(* Logix 5000 project; controller PLC_MCC1300_75F1 vendor 1 type 14 code 166 rev 32.11; software revision 32.04; part 22 of 83 *)
(* tags used below, declared in another part *)
   CM_LineToConveyorStacker_JS1 : CM_LineToConveyorStacker;
   GP_OB_InitializeMain : GP_OB_Initialize;
   M312 : MAC_Conveyor_Single;
   M312_Data : UDT_Convoy_SL;
   M312_HMW : MAC_Conveyor_HMW;
   M312_M3_ChangeSpeed : BOOL;
   M312_M3_DR_IN_MAJ : MOTION_INSTRUCTION;
   M312_M3_DR_L : AXIS_CIP_DRIVE;
   M312_M3_DR_OUT_MAJ : MOTION_INSTRUCTION;
   M312_M3_DR_OUT_MAS : MOTION_INSTRUCTION;
   M312_M3_DR_OUT_MCD : MOTION_INSTRUCTION;
   M312_SpaceConv_Utilities : SpaceConv_Utilities;
   M315_M4_DR_B1 : AXIS_CIP_DRIVE;
   M315A : MAC_Conveyor;
   M315A_ALM : MAC_Conveyor_ALM;
   M315A_Data : UDT_Convoy_SL;
   M315A_HMR : MAC_Conveyor_HMR;
   M315A_HMW : MAC_Conveyor_HMW;
   M315A_M1_DR : AXIS_CIP_DRIVE;
   M315A_M1_DR_IN_MAJ : MOTION_INSTRUCTION;
   M315A_M1_DR_IN_MAR : MOTION_INSTRUCTION;
   M315A_M1_DR_IN_MAS : MOTION_INSTRUCTION;
   M315A_M1_DR_IN_MRP : MOTION_INSTRUCTION;
   M315A_M1_DR_MAFR : MOTION_INSTRUCTION;
   M315A_M1_DR_MDR : MOTION_INSTRUCTION;
   M315A_M1_DR_MSF : MOTION_INSTRUCTION;
   M315A_M1_DR_MSO : MOTION_INSTRUCTION;
   M315A_M1_DR_OUT_MAJ : MOTION_INSTRUCTION;
   M315A_M1_DR_OUT_MAM : MOTION_INSTRUCTION;
   M315A_M1_DR_OUT_MAR : MOTION_INSTRUCTION;
   M315A_M1_DR_OUT_MAS : MOTION_INSTRUCTION;
   M315A_M1_DR_OUT_MCD : MOTION_INSTRUCTION;
   M315A_M1_DR_OUT_MRP : MOTION_INSTRUCTION;
   M315A_SpaceConv_Utilities : SpaceConv_Utilities;
   M315B : MAC_Conveyor;
   M315B_ALM : MAC_Conveyor_ALM;
   M315B_HMR : MAC_Conveyor_HMR;
   M315B_HMW : MAC_Conveyor_HMW;
   M315B_M1_DR_MAFR : MOTION_INSTRUCTION;
   M315B_M1_DR_MSF : MOTION_INSTRUCTION;
   M315B_M1_DR_MSO : MOTION_INSTRUCTION;
   M315B_M1_DR_OUT_MAR : MOTION_INSTRUCTION;
   M315B_M1_DR_OUT_MRP : MOTION_INSTRUCTION;
   M316 : MAC_Conveyor;
   TMP_dDirection : DINT;
   TMP_r : REAL;
   TMP_rAcc : REAL;
   TMP_rDec : REAL;
   TMP_rSpeed : REAL;
   TMP_rTarget_M1 : REAL;
   TMP_xForwardCommadnForCleaningZone : BOOL;
   TMP_xPositioning_M1 : BOOL;
   TMP_xPositioning_M2 : BOOL;
   TMP_xPositioning_M3 : BOOL;
   TMP_xPowerSaving : BOOL;
   TMP_xReverse_M1 : BOOL;
   TMP_xReverse_M2 : BOOL;
   TMP_xReverse_M3 : BOOL;
   TMP_xRun_M1 : BOOL;
   TMP_xRun_M2 : BOOL;
   TMP_xRun_M3 : BOOL;
   xAlwaysOFF : BOOL;
   xAlwaysON : BOOL;
   xDebugOFF : BOOL;
   Z401 : MAC_Zone;
   Z402 : MAC_Zone;
   Z402_HMW : MAC_Zone_HMW;
(* CommandLogic, continued *)

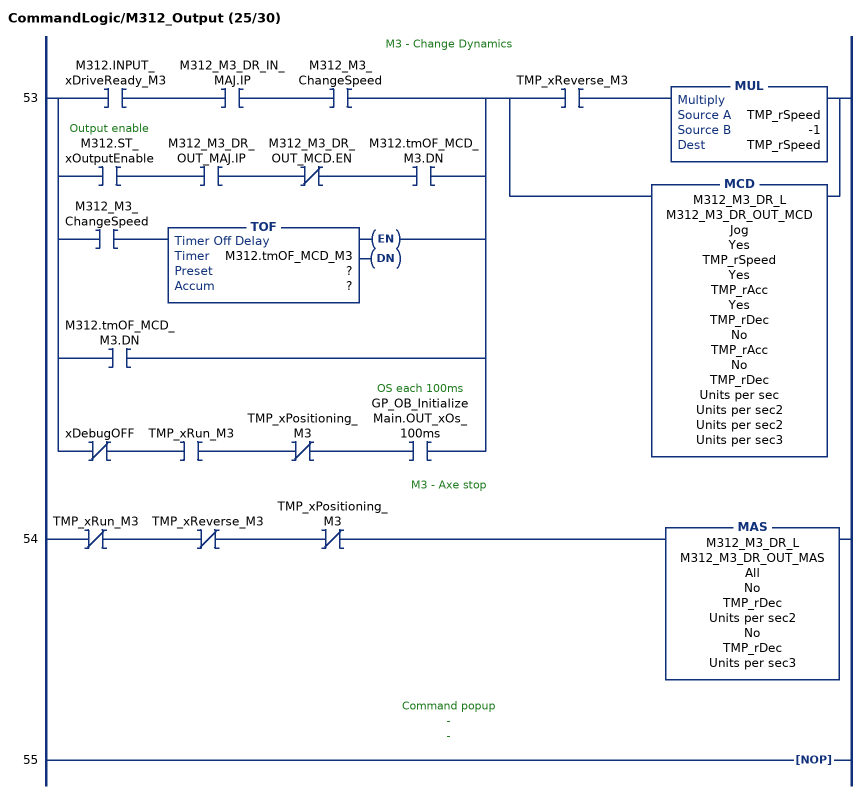
   [picture p215: CommandLogic/M312_Output rungs 53-55]
   // M3 - Change Dynamics
   53: [XIC(M312.INPUT_xDriveReady_M3) XIC(M312_M3_DR_IN_MAJ.IP) XIC(M312_M3_ChangeSpeed) ,XIC(M312.ST_xOutputEnable) XIC(M312_M3_DR_OUT_MAJ.IP) XIO(M312_M3_DR_OUT_MCD.EN) XIC(M312.tmOF_MCD_M3.DN) ,[XIC(M312_M3_ChangeSpeed) TOF(M312.tmOF_MCD_M3,?,?) ,XIC(M312.tmOF_MCD_M3.DN) ] ,XIO(xDebugOFF) XIC(TMP_xRun_M3) XIO(TMP_xPositioning_M3) XIC(GP_OB_InitializeMain.OUT_xOs_100ms) ][XIC(TMP_xReverse_M3) MUL(TMP_rSpeed,-1,TMP_rSpeed) ,MCD(M312_M3_DR_L,M312_M3_DR_OUT_MCD,Jog,Yes,TMP_rSpeed,Yes,TMP_rAcc,Yes,TMP_rDec,No,TMP_rAcc,No,TMP_rDec,Units per sec,Units per sec2,Units per sec2,Units per sec3) ];
   // M3 - Axe stop
   54: XIO(TMP_xRun_M3)XIO(TMP_xReverse_M3)XIO(TMP_xPositioning_M3)MAS(M312_M3_DR_L,M312_M3_DR_OUT_MAS,All,No,TMP_rDec,Units per sec2,No,TMP_rDec,Units per sec3);
   // Command popup
   // -
   // -
   55: NOP();
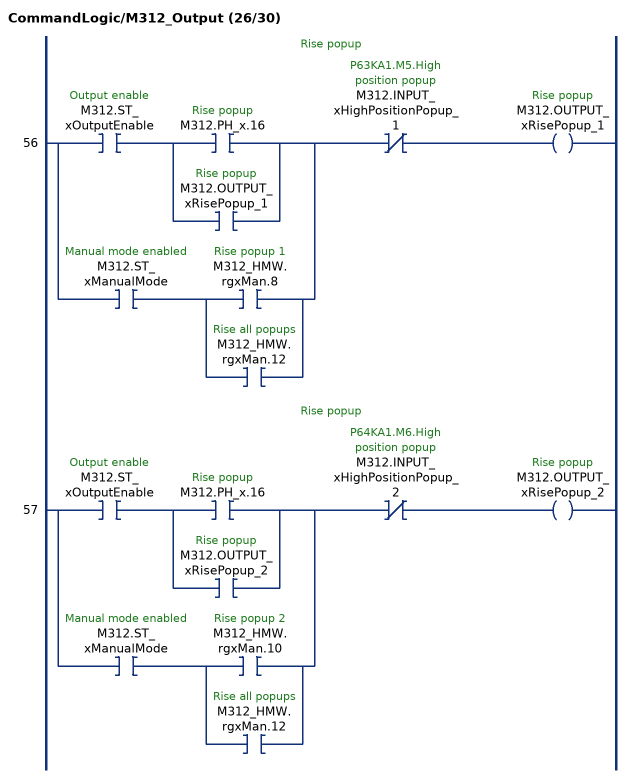
   // Rise popup
   56: [XIC(M312.ST_xOutputEnable) [XIC(M312.PH_x.16) ,XIC(M312.OUTPUT_xRisePopup_1) ] ,XIC(M312.ST_xManualMode) [XIC(M312_HMW.rgxMan.8) ,XIC(M312_HMW.rgxMan.12) ] ]XIO(M312.INPUT_xHighPositionPopup_1)OTE(M312.OUTPUT_xRisePopup_1);
   // Rise popup
   57: [XIC(M312.ST_xOutputEnable) [XIC(M312.PH_x.16) ,XIC(M312.OUTPUT_xRisePopup_2) ] ,XIC(M312.ST_xManualMode) [XIC(M312_HMW.rgxMan.10) ,XIC(M312_HMW.rgxMan.12) ] ]XIO(M312.INPUT_xHighPositionPopup_2)OTE(M312.OUTPUT_xRisePopup_2);
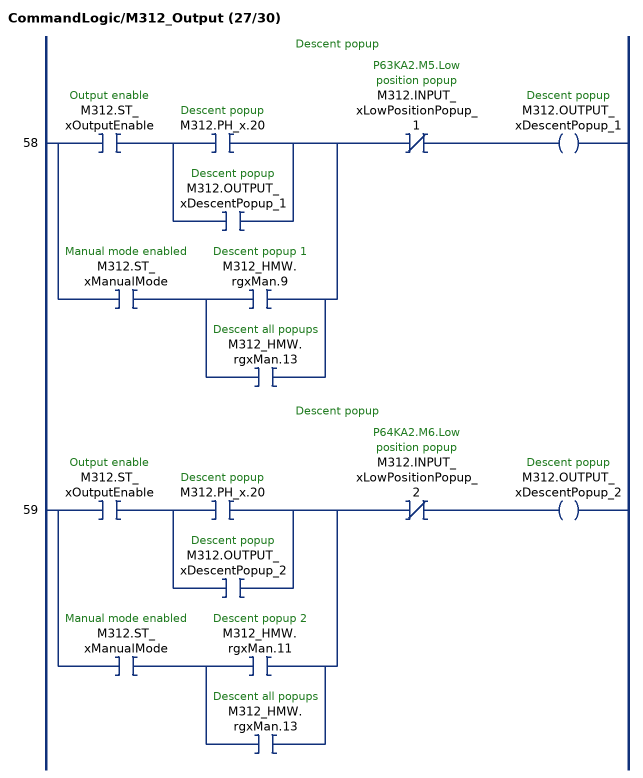
   // Descent popup
   58: [XIC(M312.ST_xOutputEnable) [XIC(M312.PH_x.20) ,XIC(M312.OUTPUT_xDescentPopup_1) ] ,XIC(M312.ST_xManualMode) [XIC(M312_HMW.rgxMan.9) ,XIC(M312_HMW.rgxMan.13) ] ]XIO(M312.INPUT_xLowPositionPopup_1)OTE(M312.OUTPUT_xDescentPopup_1);
   // Descent popup
   59: [XIC(M312.ST_xOutputEnable) [XIC(M312.PH_x.20) ,XIC(M312.OUTPUT_xDescentPopup_2) ] ,XIC(M312.ST_xManualMode) [XIC(M312_HMW.rgxMan.11) ,XIC(M312_HMW.rgxMan.13) ] ]XIO(M312.INPUT_xLowPositionPopup_2)OTE(M312.OUTPUT_xDescentPopup_2);
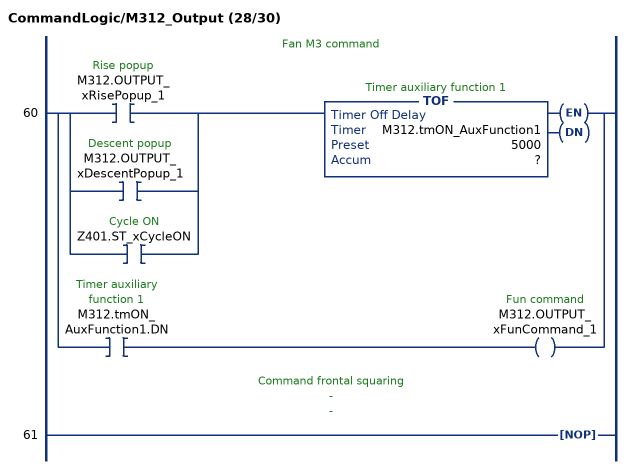
   // Fan M3 command
   60: [[XIC(M312.OUTPUT_xRisePopup_1) ,[XIC(M312.OUTPUT_xDescentPopup_1) ,XIC(Z401.ST_xCycleON) ] ] TOF(M312.tmON_AuxFunction1,?,?) ,XIC(M312.tmON_AuxFunction1.DN) OTE(M312.OUTPUT_xFunCommand_1) ];
   // Command frontal squaring
   // -
   // -
   61: NOP();
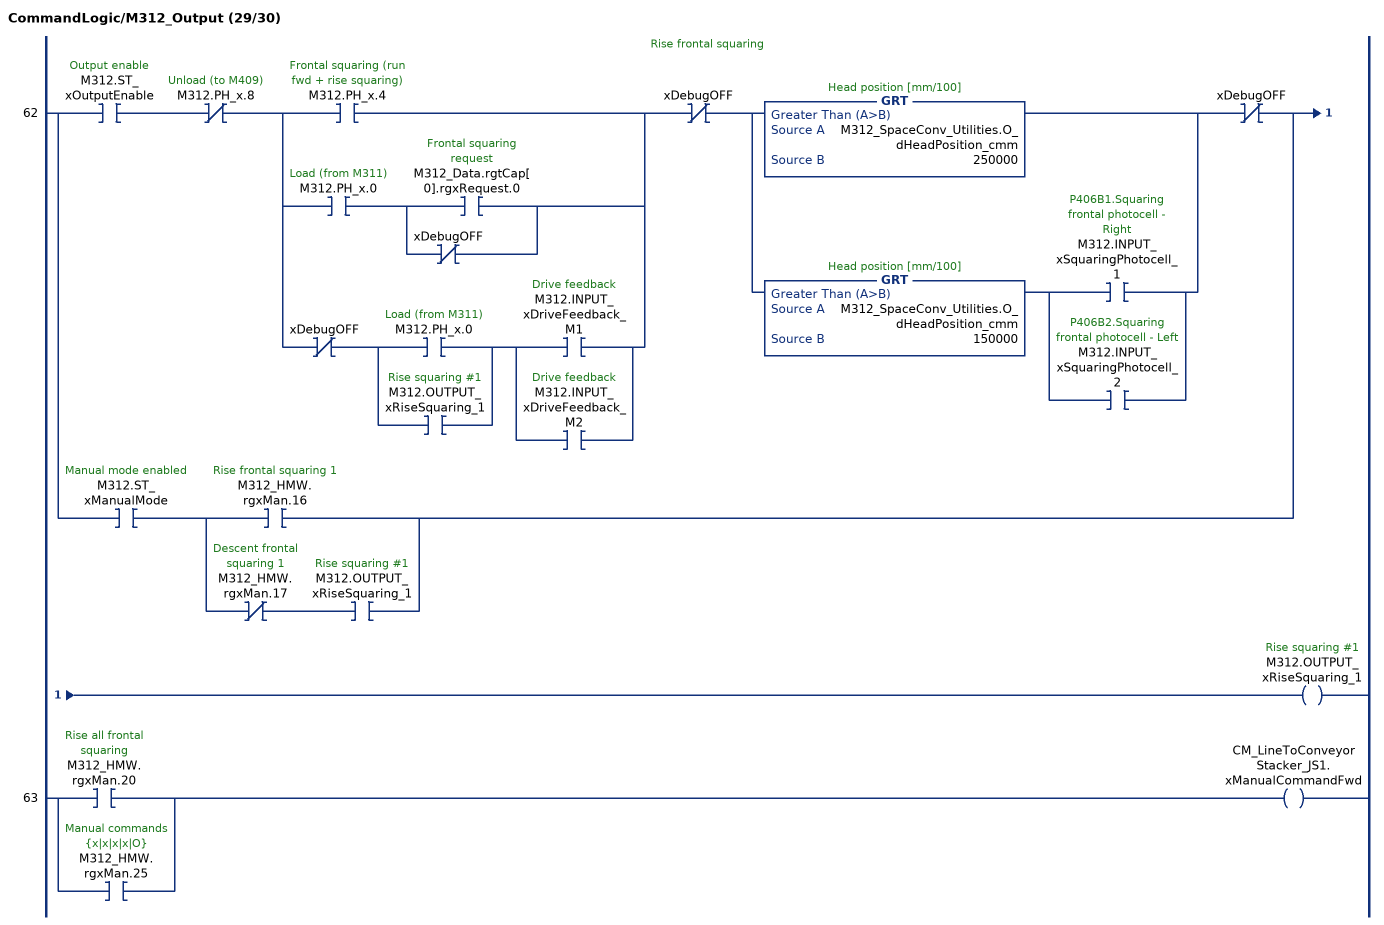
   // Rise frontal squaring
   62: [XIC(M312.ST_xOutputEnable) XIO(M312.PH_x.8) [XIC(M312.PH_x.4) ,XIC(M312.PH_x.0) [XIC(M312_Data.rgtCap[0].rgxRequest.0) ,XIO(xDebugOFF) ] ,XIO(xDebugOFF) [XIC(M312.PH_x.0) ,XIC(M312.OUTPUT_xRiseSquaring_1) ] [XIC(M312.INPUT_xDriveFeedback_M1) ,XIC(M312.INPUT_xDriveFeedback_M2) ] ] XIO(xDebugOFF) [GRT(M312_SpaceConv_Utilities.O_dHeadPosition_cmm,250000) ,GRT(M312_SpaceConv_Utilities.O_dHeadPosition_cmm,150000) [XIC(M312.INPUT_xSquaringPhotocell_1) ,XIC(M312.INPUT_xSquaringPhotocell_2) ] ] XIO(xDebugOFF) ,XIC(M312.ST_xManualMode) [XIC(M312_HMW.rgxMan.16) ,XIO(M312_HMW.rgxMan.17) XIC(M312.OUTPUT_xRiseSquaring_1) ] ]OTE(M312.OUTPUT_xRiseSquaring_1);
   63: [XIC(M312_HMW.rgxMan.20) ,XIC(M312_HMW.rgxMan.25) ]OTE(CM_LineToConveyorStacker_JS1.xManualCommandFwd);
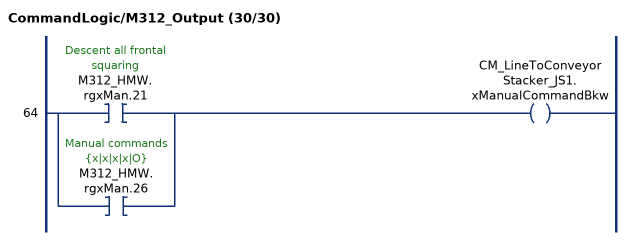
   64: [XIC(M312_HMW.rgxMan.21) ,XIC(M312_HMW.rgxMan.26) ]OTE(CM_LineToConveyorStacker_JS1.xManualCommandBkw);
END_ROUTINE

ROUTINE M315A_Output   (* ladder *)
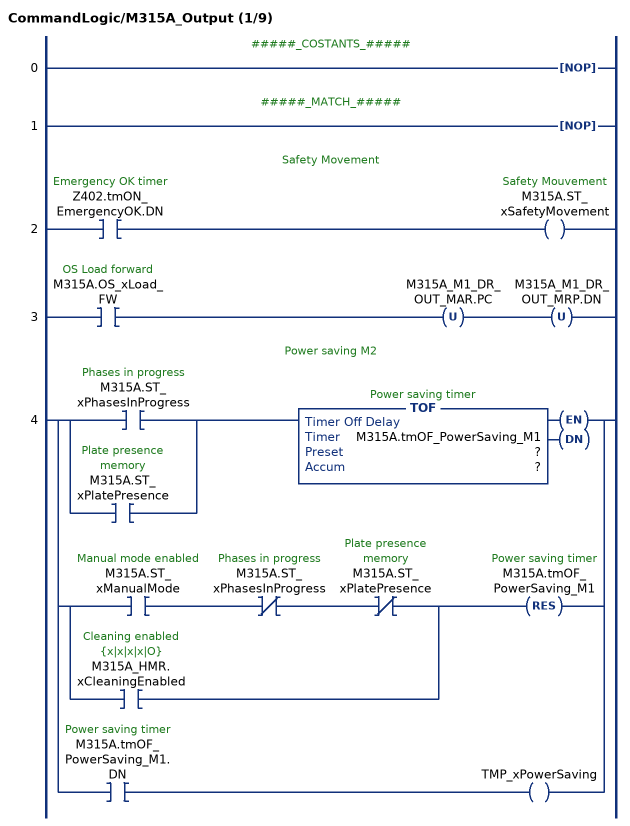
   // #####_COSTANTS_#####
   0: NOP();
   // #####_MATCH_#####
   1: NOP();
   // Safety Movement
   2: XIC(Z402.tmON_EmergencyOK.DN)OTE(M315A.ST_xSafetyMovement);
   3: XIC(M315A.OS_xLoad_FW)OTU(M315A_M1_DR_OUT_MAR.PC)OTU(M315A_M1_DR_OUT_MRP.DN);
   // Power saving M2
   4: [[XIC(M315A.ST_xPhasesInProgress) ,XIC(M315A.ST_xPlatePresence) ] TOF(M315A.tmOF_PowerSaving_M1,?,?) ,[XIC(M315A.ST_xManualMode) XIO(M315A.ST_xPhasesInProgress) XIO(M315A.ST_xPlatePresence) ,XIC(M315A_HMR.xCleaningEnabled) ] RES(M315A.tmOF_PowerSaving_M1) ,XIC(M315A.tmOF_PowerSaving_M1.DN) OTE(TMP_xPowerSaving) ];
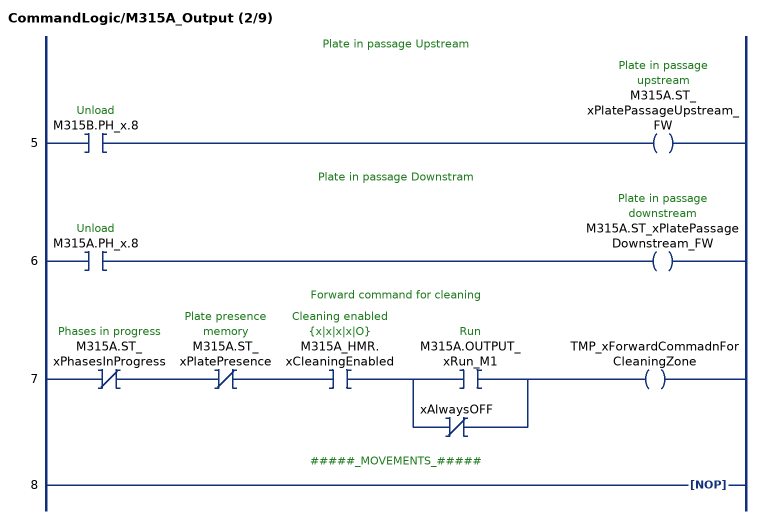
   // Plate in passage Upstream
   5: XIC(M315B.PH_x.8)OTE(M315A.ST_xPlatePassageUpstream_FW);
   // Plate in passage Downstram
   6: XIC(M315A.PH_x.8)OTE(M315A.ST_xPlatePassageDownstream_FW);
   // Forward command for cleaning
   7: XIO(M315A.ST_xPhasesInProgress)XIO(M315A.ST_xPlatePresence)XIC(M315A_HMR.xCleaningEnabled)[XIC(M315A.OUTPUT_xRun_M1) ,XIO(xAlwaysOFF) ]OTE(TMP_xForwardCommadnForCleaningZone);
   // #####_MOVEMENTS_#####
   8: NOP();
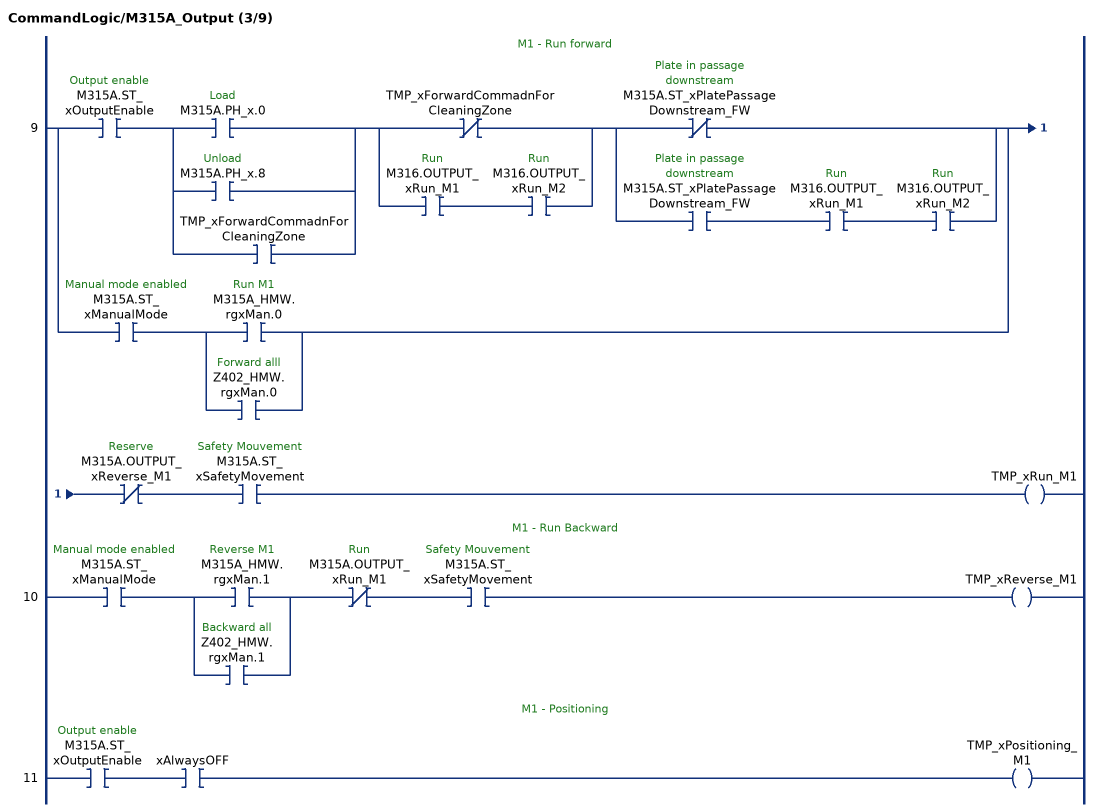
   // M1 - Run forward
   9: [XIC(M315A.ST_xOutputEnable) [XIC(M315A.PH_x.0) ,XIC(M315A.PH_x.8) ,XIC(TMP_xForwardCommadnForCleaningZone) ] [XIO(TMP_xForwardCommadnForCleaningZone) ,XIC(M316.OUTPUT_xRun_M1) XIC(M316.OUTPUT_xRun_M2) ] [XIO(M315A.ST_xPlatePassageDownstream_FW) ,XIC(M315A.ST_xPlatePassageDownstream_FW) XIC(M316.OUTPUT_xRun_M1) XIC(M316.OUTPUT_xRun_M2) ] ,XIC(M315A.ST_xManualMode) [XIC(M315A_HMW.rgxMan.0) ,XIC(Z402_HMW.rgxMan.0) ] ]XIO(M315A.OUTPUT_xReverse_M1)XIC(M315A.ST_xSafetyMovement)OTE(TMP_xRun_M1);
   // M1 - Run Backward
   10: XIC(M315A.ST_xManualMode)[XIC(M315A_HMW.rgxMan.1) ,XIC(Z402_HMW.rgxMan.1) ]XIO(M315A.OUTPUT_xRun_M1)XIC(M315A.ST_xSafetyMovement)OTE(TMP_xReverse_M1);
   // M1 - Positioning
   11: XIC(M315A.ST_xOutputEnable)XIC(xAlwaysOFF)OTE(TMP_xPositioning_M1);
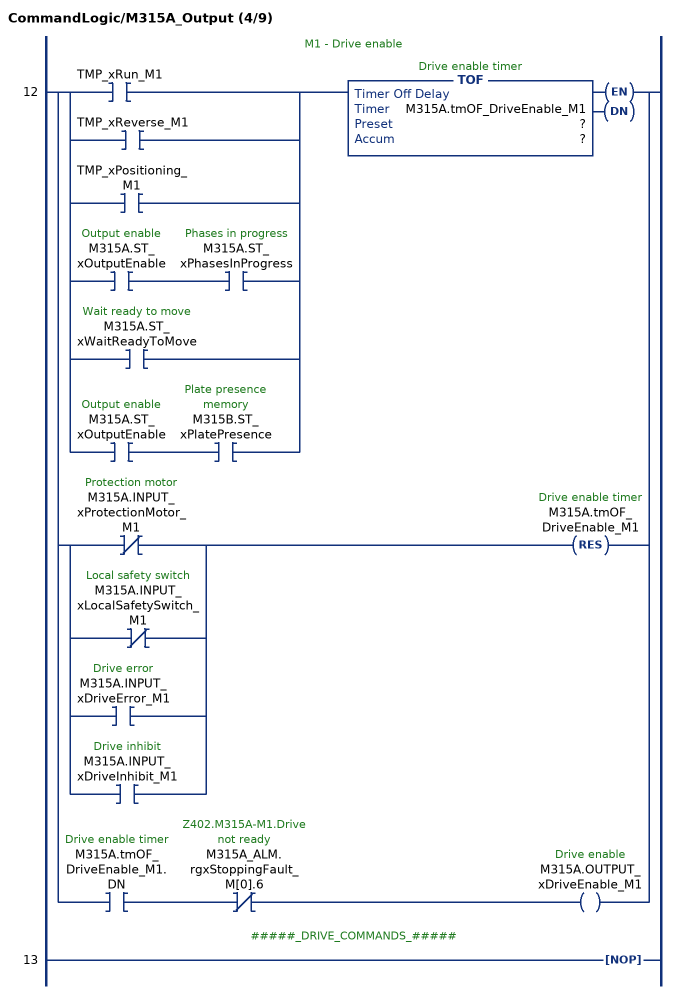
   // M1 - Drive enable
   12: [[XIC(TMP_xRun_M1) ,XIC(TMP_xReverse_M1) ,XIC(TMP_xPositioning_M1) ,XIC(M315A.ST_xOutputEnable) XIC(M315A.ST_xPhasesInProgress) ,XIC(M315A.ST_xWaitReadyToMove) ,XIC(M315A.ST_xOutputEnable) XIC(M315B.ST_xPlatePresence) ] TOF(M315A.tmOF_DriveEnable_M1,?,?) ,[XIO(M315A.INPUT_xProtectionMotor_M1) ,XIO(M315A.INPUT_xLocalSafetySwitch_M1) ,XIC(M315A.INPUT_xDriveError_M1) ,XIC(M315A.INPUT_xDriveInhibit_M1) ] RES(M315A.tmOF_DriveEnable_M1) ,XIC(M315A.tmOF_DriveEnable_M1.DN) XIO(M315A_ALM.rgxStoppingFault_M[0].6) OTE(M315A.OUTPUT_xDriveEnable_M1) ];
   // #####_DRIVE_COMMANDS_#####
   13: NOP();
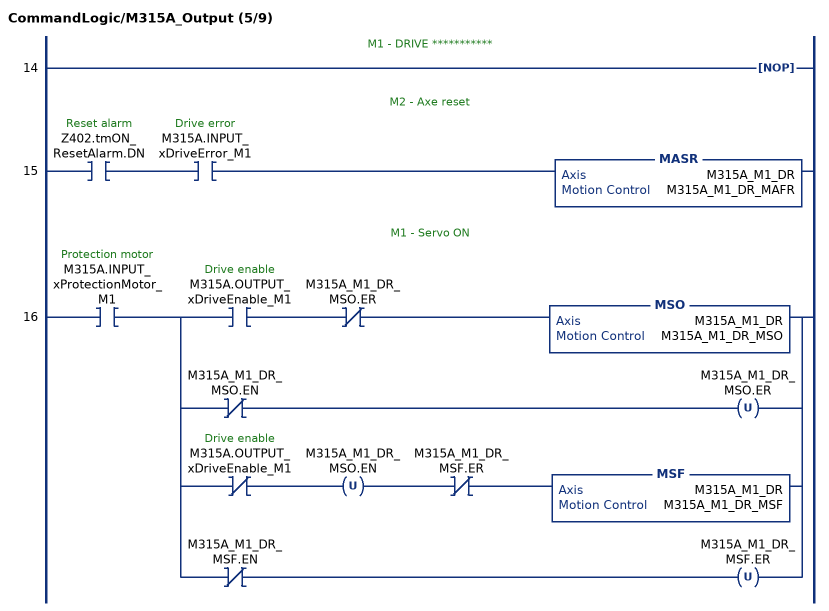
   // M1 - DRIVE ***********
   14: NOP();
   // M2 - Axe reset
   15: XIC(Z402.tmON_ResetAlarm.DN)XIC(M315A.INPUT_xDriveError_M1)MASR(M315A_M1_DR,M315A_M1_DR_MAFR);
   // M1 - Servo ON
   16: XIC(M315A.INPUT_xProtectionMotor_M1)[XIC(M315A.OUTPUT_xDriveEnable_M1) XIO(M315A_M1_DR_MSO.ER) MSO(M315A_M1_DR,M315A_M1_DR_MSO) ,XIO(M315A_M1_DR_MSO.EN) OTU(M315A_M1_DR_MSO.ER) ,XIO(M315A.OUTPUT_xDriveEnable_M1) OTU(M315A_M1_DR_MSO.EN) XIO(M315A_M1_DR_MSF.ER) MSF(M315A_M1_DR,M315A_M1_DR_MSF) ,XIO(M315A_M1_DR_MSF.EN) OTU(M315A_M1_DR_MSF.ER) ];
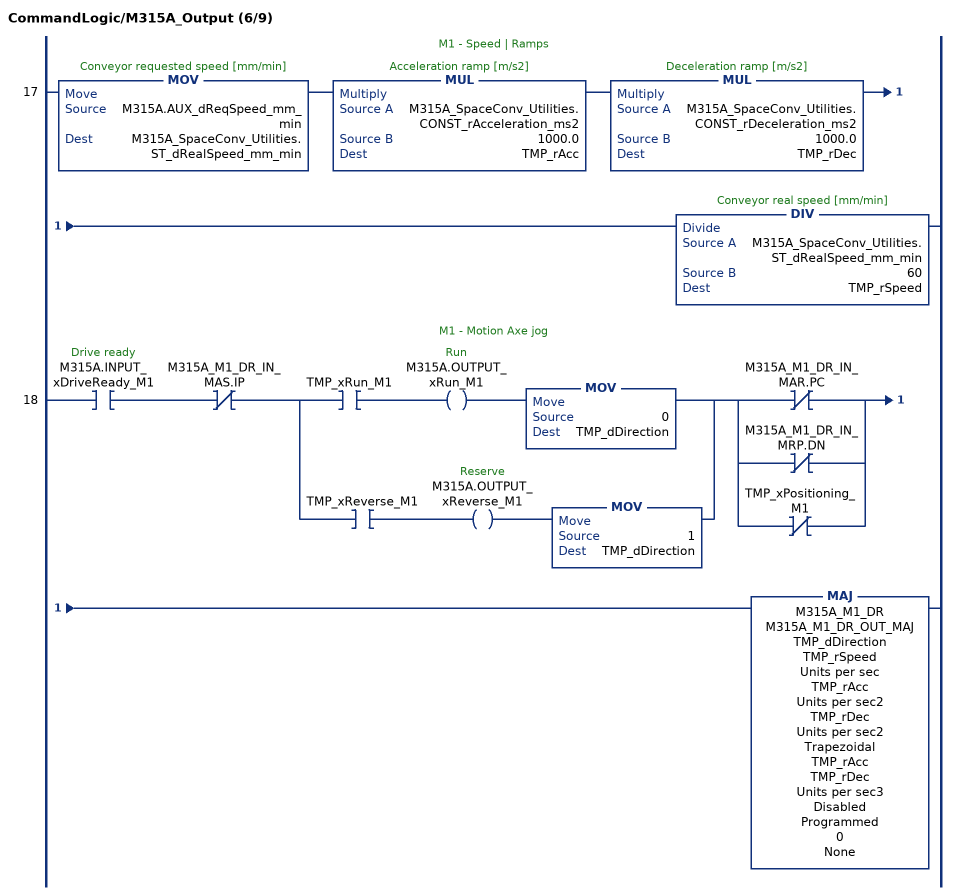
   // M1 - Speed | Ramps
   17: MOV(M315A.AUX_dReqSpeed_mm_min,M315A_SpaceConv_Utilities.ST_dRealSpeed_mm_min)MUL(M315A_SpaceConv_Utilities.CONST_rAcceleration_ms2,1000.0,TMP_rAcc)MUL(M315A_SpaceConv_Utilities.CONST_rDeceleration_ms2,1000.0,TMP_rDec)DIV(M315A_SpaceConv_Utilities.ST_dRealSpeed_mm_min,60,TMP_rSpeed);
   // M1 - Motion Axe jog
   18: XIC(M315A.INPUT_xDriveReady_M1)XIO(M315A_M1_DR_IN_MAS.IP)[XIC(TMP_xRun_M1) OTE(M315A.OUTPUT_xRun_M1) MOV(0,TMP_dDirection) ,XIC(TMP_xReverse_M1) OTE(M315A.OUTPUT_xReverse_M1) MOV(1,TMP_dDirection) ][XIO(M315A_M1_DR_IN_MAR.PC) ,XIO(M315A_M1_DR_IN_MRP.DN) ,XIO(TMP_xPositioning_M1) ]MAJ(M315A_M1_DR,M315A_M1_DR_OUT_MAJ,TMP_dDirection,TMP_rSpeed,Units per sec,TMP_rAcc,Units per sec2,TMP_rDec,Units per sec2,Trapezoidal,TMP_rAcc,TMP_rDec,Units per sec3,Disabled,Programmed,0,None);
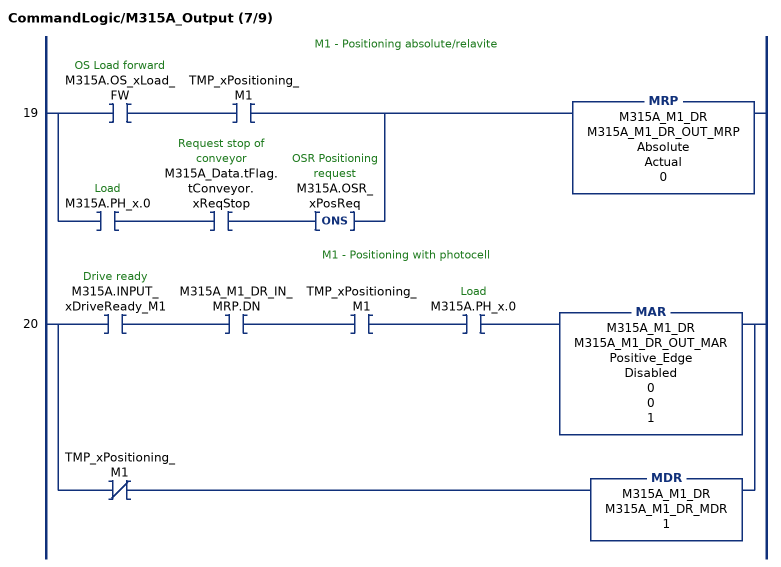
   // M1 - Positioning absolute/relavite
   19: [XIC(M315A.OS_xLoad_FW) XIC(TMP_xPositioning_M1) ,XIC(M315A.PH_x.0) XIC(M315A_Data.tFlag.tConveyor.xReqStop) ONS(M315A.OSR_xPosReq) ]MRP(M315A_M1_DR,M315A_M1_DR_OUT_MRP,Absolute,Actual,0);
   // M1 - Positioning with photocell
   20: [XIC(M315A.INPUT_xDriveReady_M1) XIC(M315A_M1_DR_IN_MRP.DN) XIC(TMP_xPositioning_M1) XIC(M315A.PH_x.0) MAR(M315A_M1_DR,M315A_M1_DR_OUT_MAR,Positive_Edge,Disabled,0,0,1) ,XIO(TMP_xPositioning_M1) MDR(M315A_M1_DR,M315A_M1_DR_MDR,1) ];
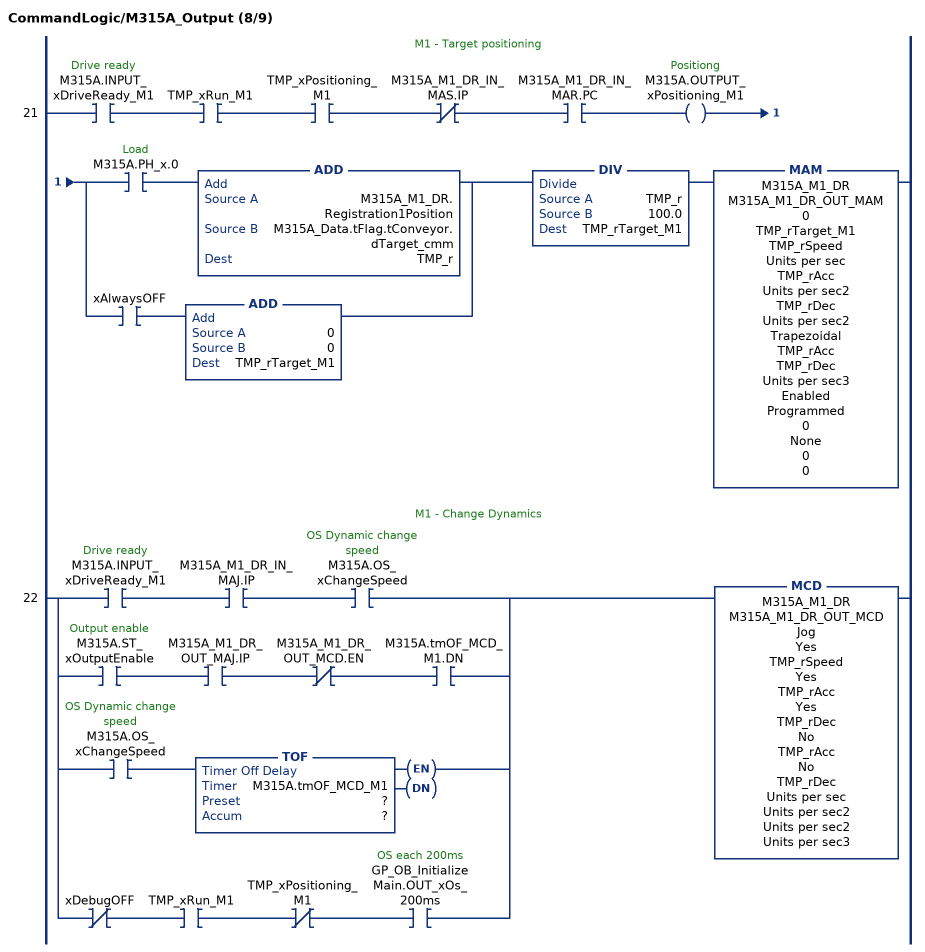
   // M1 - Target positioning
   21: XIC(M315A.INPUT_xDriveReady_M1)XIC(TMP_xRun_M1)XIC(TMP_xPositioning_M1)XIO(M315A_M1_DR_IN_MAS.IP)XIC(M315A_M1_DR_IN_MAR.PC)OTE(M315A.OUTPUT_xPositioning_M1)[XIC(M315A.PH_x.0) ADD(M315A_M1_DR.Registration1Position,M315A_Data.tFlag.tConveyor.dTarget_cmm,TMP_r) ,XIC(xAlwaysOFF) ADD(0,0,TMP_rTarget_M1) ]DIV(TMP_r,100.0,TMP_rTarget_M1)MAM(M315A_M1_DR,M315A_M1_DR_OUT_MAM,0,TMP_rTarget_M1,TMP_rSpeed,Units per sec,TMP_rAcc,Units per sec2,TMP_rDec,Units per sec2,Trapezoidal,TMP_rAcc,TMP_rDec,Units per sec3,Enabled,Programmed,0,None,0,0);
   // M1 - Change Dynamics
   22: [XIC(M315A.INPUT_xDriveReady_M1) XIC(M315A_M1_DR_IN_MAJ.IP) XIC(M315A.OS_xChangeSpeed) ,XIC(M315A.ST_xOutputEnable) XIC(M315A_M1_DR_OUT_MAJ.IP) XIO(M315A_M1_DR_OUT_MCD.EN) XIC(M315A.tmOF_MCD_M1.DN) ,XIC(M315A.OS_xChangeSpeed) TOF(M315A.tmOF_MCD_M1,?,?) ,XIO(xDebugOFF) XIC(TMP_xRun_M1) XIO(TMP_xPositioning_M1) XIC(GP_OB_InitializeMain.OUT_xOs_200ms) ]MCD(M315A_M1_DR,M315A_M1_DR_OUT_MCD,Jog,Yes,TMP_rSpeed,Yes,TMP_rAcc,Yes,TMP_rDec,No,TMP_rAcc,No,TMP_rDec,Units per sec,Units per sec2,Units per sec2,Units per sec3);
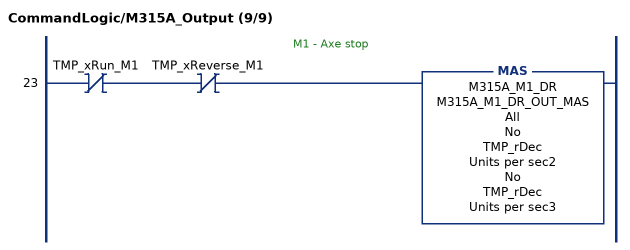
   // M1 - Axe stop
   23: XIO(TMP_xRun_M1)XIO(TMP_xReverse_M1)MAS(M315A_M1_DR,M315A_M1_DR_OUT_MAS,All,No,TMP_rDec,Units per sec2,No,TMP_rDec,Units per sec3);
END_ROUTINE

ROUTINE M315B_Output   (* ladder *)
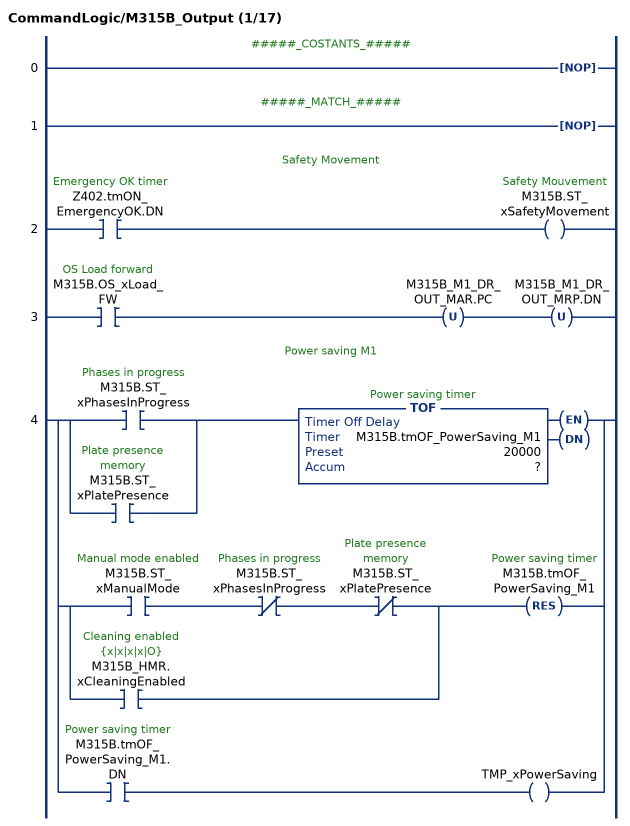
   // #####_COSTANTS_#####
   0: NOP();
   // #####_MATCH_#####
   1: NOP();
   // Safety Movement
   2: XIC(Z402.tmON_EmergencyOK.DN)OTE(M315B.ST_xSafetyMovement);
   3: XIC(M315B.OS_xLoad_FW)OTU(M315B_M1_DR_OUT_MAR.PC)OTU(M315B_M1_DR_OUT_MRP.DN);
   // Power saving M1
   4: [[XIC(M315B.ST_xPhasesInProgress) ,XIC(M315B.ST_xPlatePresence) ] TOF(M315B.tmOF_PowerSaving_M1,?,?) ,[XIC(M315B.ST_xManualMode) XIO(M315B.ST_xPhasesInProgress) XIO(M315B.ST_xPlatePresence) ,XIC(M315B_HMR.xCleaningEnabled) ] RES(M315B.tmOF_PowerSaving_M1) ,XIC(M315B.tmOF_PowerSaving_M1.DN) OTE(TMP_xPowerSaving) ];
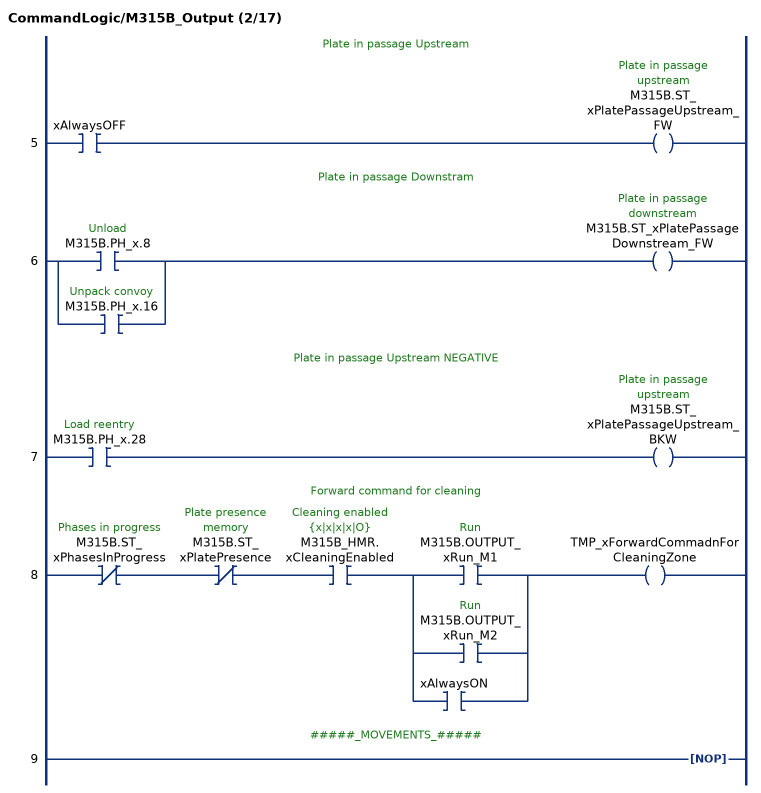
   // Plate in passage Upstream
   5: XIC(xAlwaysOFF)OTE(M315B.ST_xPlatePassageUpstream_FW);
   // Plate in passage Downstram
   6: [XIC(M315B.PH_x.8) ,XIC(M315B.PH_x.16) ]OTE(M315B.ST_xPlatePassageDownstream_FW);
   // Plate in passage Upstream NEGATIVE
   7: XIC(M315B.PH_x.28)OTE(M315B.ST_xPlatePassageUpstream_BKW);
   // Forward command for cleaning
   8: XIO(M315B.ST_xPhasesInProgress)XIO(M315B.ST_xPlatePresence)XIC(M315B_HMR.xCleaningEnabled)[XIC(M315B.OUTPUT_xRun_M1) ,XIC(M315B.OUTPUT_xRun_M2) ,XIC(xAlwaysON) ]OTE(TMP_xForwardCommadnForCleaningZone);
   // #####_MOVEMENTS_#####
   9: NOP();
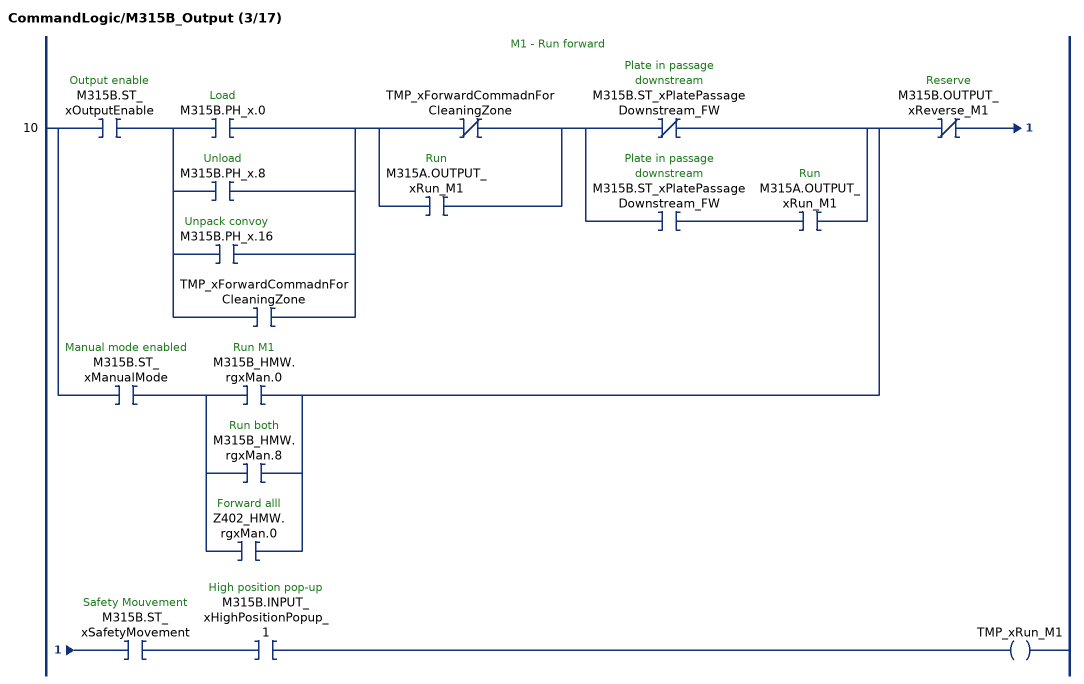
   // M1 - Run forward
   10: [XIC(M315B.ST_xOutputEnable) [XIC(M315B.PH_x.0) ,XIC(M315B.PH_x.8) ,XIC(M315B.PH_x.16) ,XIC(TMP_xForwardCommadnForCleaningZone) ] [XIO(TMP_xForwardCommadnForCleaningZone) ,XIC(M315A.OUTPUT_xRun_M1) ] [XIO(M315B.ST_xPlatePassageDownstream_FW) ,XIC(M315B.ST_xPlatePassageDownstream_FW) XIC(M315A.OUTPUT_xRun_M1) ] ,XIC(M315B.ST_xManualMode) [XIC(M315B_HMW.rgxMan.0) ,XIC(M315B_HMW.rgxMan.8) ,XIC(Z402_HMW.rgxMan.0) ] ]XIO(M315B.OUTPUT_xReverse_M1)XIC(M315B.ST_xSafetyMovement)XIC(M315B.INPUT_xHighPositionPopup_1)OTE(TMP_xRun_M1);
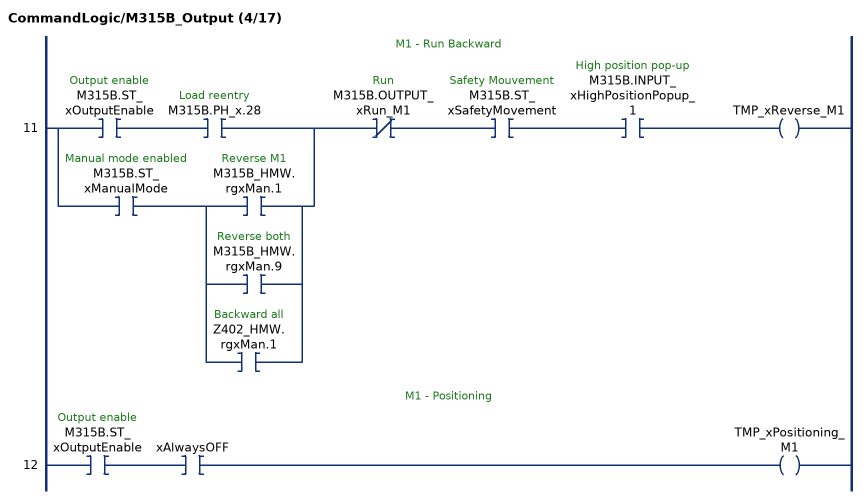
   // M1 - Run Backward
   11: [XIC(M315B.ST_xOutputEnable) XIC(M315B.PH_x.28) ,XIC(M315B.ST_xManualMode) [XIC(M315B_HMW.rgxMan.1) ,XIC(M315B_HMW.rgxMan.9) ,XIC(Z402_HMW.rgxMan.1) ] ]XIO(M315B.OUTPUT_xRun_M1)XIC(M315B.ST_xSafetyMovement)XIC(M315B.INPUT_xHighPositionPopup_1)OTE(TMP_xReverse_M1);
   // M1 - Positioning
   12: XIC(M315B.ST_xOutputEnable)XIC(xAlwaysOFF)OTE(TMP_xPositioning_M1);
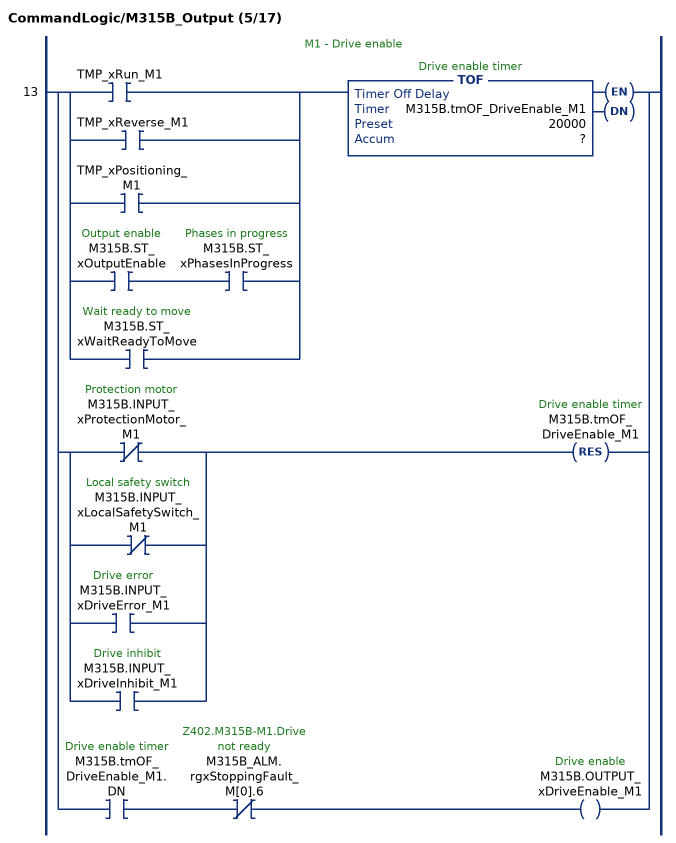
   // M1 - Drive enable
   13: [[XIC(TMP_xRun_M1) ,XIC(TMP_xReverse_M1) ,XIC(TMP_xPositioning_M1) ,XIC(M315B.ST_xOutputEnable) XIC(M315B.ST_xPhasesInProgress) ,XIC(M315B.ST_xWaitReadyToMove) ] TOF(M315B.tmOF_DriveEnable_M1,?,?) ,[XIO(M315B.INPUT_xProtectionMotor_M1) ,XIO(M315B.INPUT_xLocalSafetySwitch_M1) ,XIC(M315B.INPUT_xDriveError_M1) ,XIC(M315B.INPUT_xDriveInhibit_M1) ] RES(M315B.tmOF_DriveEnable_M1) ,XIC(M315B.tmOF_DriveEnable_M1.DN) XIO(M315B_ALM.rgxStoppingFault_M[0].6) OTE(M315B.OUTPUT_xDriveEnable_M1) ];
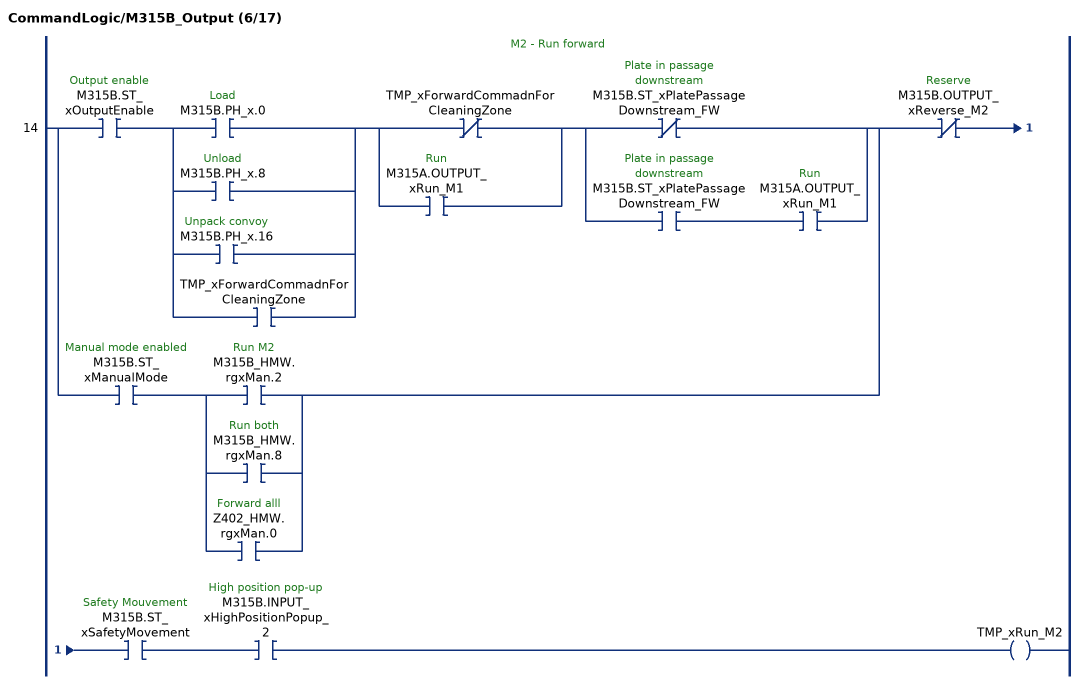
   // M2 - Run forward
   14: [XIC(M315B.ST_xOutputEnable) [XIC(M315B.PH_x.0) ,XIC(M315B.PH_x.8) ,XIC(M315B.PH_x.16) ,XIC(TMP_xForwardCommadnForCleaningZone) ] [XIO(TMP_xForwardCommadnForCleaningZone) ,XIC(M315A.OUTPUT_xRun_M1) ] [XIO(M315B.ST_xPlatePassageDownstream_FW) ,XIC(M315B.ST_xPlatePassageDownstream_FW) XIC(M315A.OUTPUT_xRun_M1) ] ,XIC(M315B.ST_xManualMode) [XIC(M315B_HMW.rgxMan.2) ,XIC(M315B_HMW.rgxMan.8) ,XIC(Z402_HMW.rgxMan.0) ] ]XIO(M315B.OUTPUT_xReverse_M2)XIC(M315B.ST_xSafetyMovement)XIC(M315B.INPUT_xHighPositionPopup_2)OTE(TMP_xRun_M2);
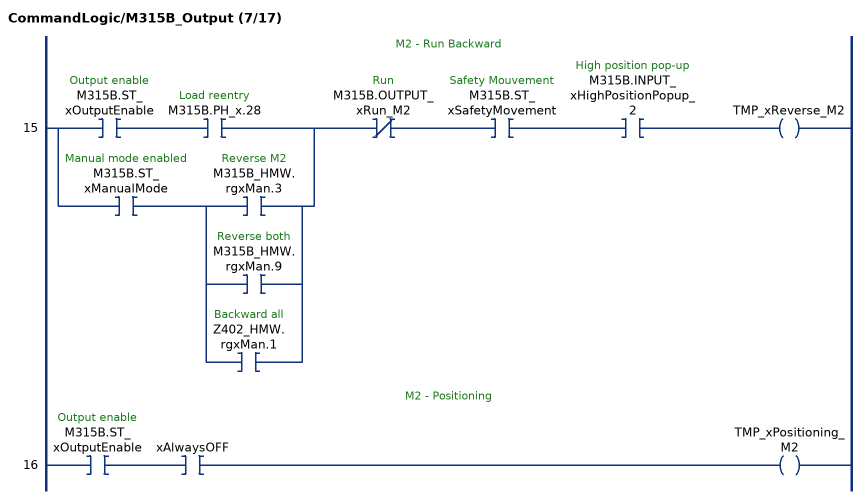
   // M2 - Run Backward
   15: [XIC(M315B.ST_xOutputEnable) XIC(M315B.PH_x.28) ,XIC(M315B.ST_xManualMode) [XIC(M315B_HMW.rgxMan.3) ,XIC(M315B_HMW.rgxMan.9) ,XIC(Z402_HMW.rgxMan.1) ] ]XIO(M315B.OUTPUT_xRun_M2)XIC(M315B.ST_xSafetyMovement)XIC(M315B.INPUT_xHighPositionPopup_2)OTE(TMP_xReverse_M2);
   // M2 - Positioning
   16: XIC(M315B.ST_xOutputEnable)XIC(xAlwaysOFF)OTE(TMP_xPositioning_M2);
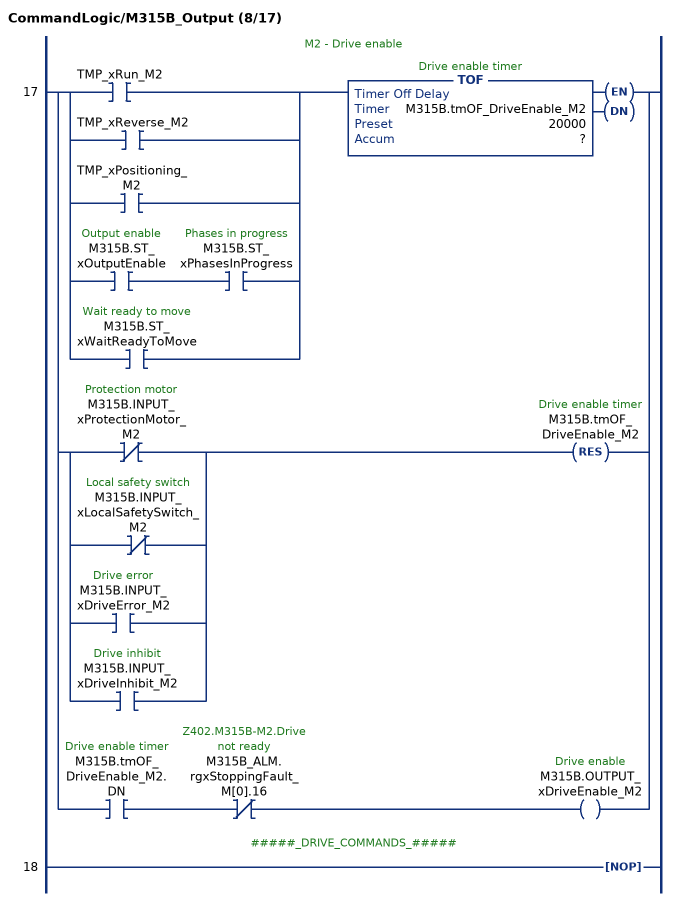
   // M2 - Drive enable
   17: [[XIC(TMP_xRun_M2) ,XIC(TMP_xReverse_M2) ,XIC(TMP_xPositioning_M2) ,XIC(M315B.ST_xOutputEnable) XIC(M315B.ST_xPhasesInProgress) ,XIC(M315B.ST_xWaitReadyToMove) ] TOF(M315B.tmOF_DriveEnable_M2,?,?) ,[XIO(M315B.INPUT_xProtectionMotor_M2) ,XIO(M315B.INPUT_xLocalSafetySwitch_M2) ,XIC(M315B.INPUT_xDriveError_M2) ,XIC(M315B.INPUT_xDriveInhibit_M2) ] RES(M315B.tmOF_DriveEnable_M2) ,XIC(M315B.tmOF_DriveEnable_M2.DN) XIO(M315B_ALM.rgxStoppingFault_M[0].16) OTE(M315B.OUTPUT_xDriveEnable_M2) ];
   // #####_DRIVE_COMMANDS_#####
   18: NOP();
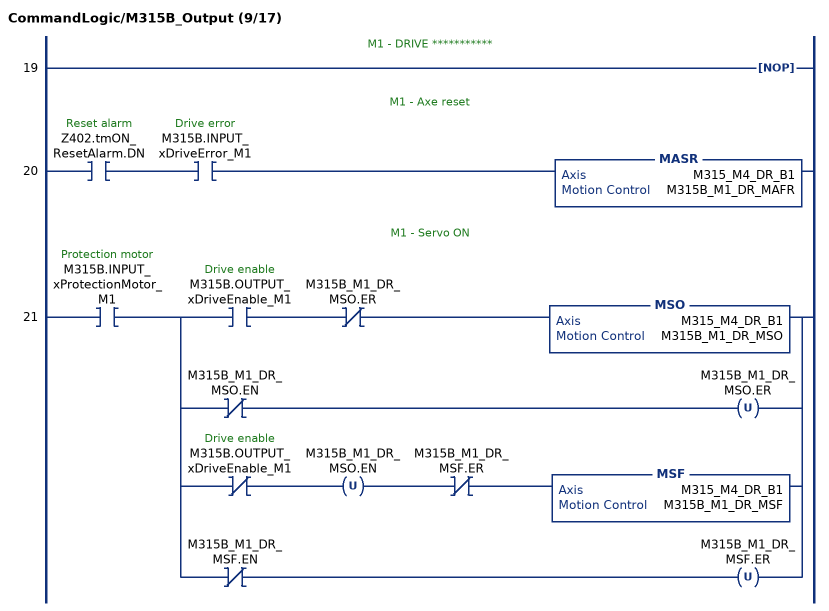
   // M1 - DRIVE ***********
   19: NOP();
   // M1 - Axe reset
   20: XIC(Z402.tmON_ResetAlarm.DN)XIC(M315B.INPUT_xDriveError_M1)MASR(M315_M4_DR_B1,M315B_M1_DR_MAFR);
   // M1 - Servo ON
   21: XIC(M315B.INPUT_xProtectionMotor_M1)[XIC(M315B.OUTPUT_xDriveEnable_M1) XIO(M315B_M1_DR_MSO.ER) MSO(M315_M4_DR_B1,M315B_M1_DR_MSO) ,XIO(M315B_M1_DR_MSO.EN) OTU(M315B_M1_DR_MSO.ER) ,XIO(M315B.OUTPUT_xDriveEnable_M1) OTU(M315B_M1_DR_MSO.EN) XIO(M315B_M1_DR_MSF.ER) MSF(M315_M4_DR_B1,M315B_M1_DR_MSF) ,XIO(M315B_M1_DR_MSF.EN) OTU(M315B_M1_DR_MSF.ER) ];
